REGION Network 93: Proximo Mantenimiento #1 MC060
   RUNG wire#powerrail
      { S7_Templates := "SrcType := DInt"; S7_GenerateENO := "TRUE" } Add(in1 := "Varios".UltimoMantMC060_1, in2 := "Varios".HorasMantMC060_1, out => "ProxMantMC060_1")
   END_RUNG
   // the same network as SCL:
   "ProxMantMC060_1" := "Varios".UltimoMantMC060_1 + "Varios".HorasMantMC060_1;
END_REGION

REGION Network 94: Se superaron las horas para el mantenimiento #1 MC060 / Animación Horas MAX Compresor de Alta ABC5
   RUNG wire#powerrail
      { S7_Templates := "SrcType := DInt" } GE_Contact(in1 := "HorasCmpBaja".HMMC060, in2 := "ProxMantMC060_1")
      Coil( "LimiteMantMC060_1" )
   END_RUNG
   // the same network as SCL:
   "LimiteMantMC060_1" := "HorasCmpBaja".HMMC060 >= "ProxMantMC060_1";
END_REGION

REGION Network 95: Proximo Mantenimiento #2 MC060
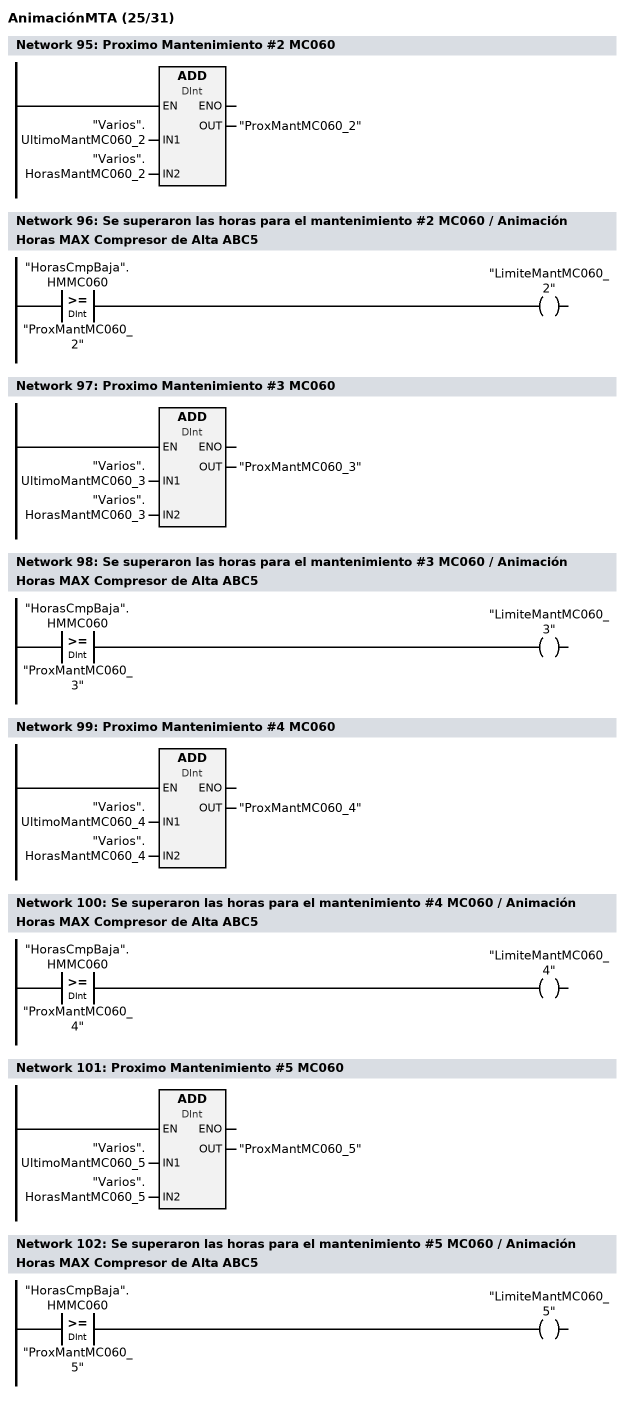
   RUNG wire#powerrail
      { S7_Templates := "SrcType := DInt"; S7_GenerateENO := "TRUE" } Add(in1 := "Varios".UltimoMantMC060_2, in2 := "Varios".HorasMantMC060_2, out => "ProxMantMC060_2")
   END_RUNG
   // the same network as SCL:
   "ProxMantMC060_2" := "Varios".UltimoMantMC060_2 + "Varios".HorasMantMC060_2;
END_REGION

REGION Network 96: Se superaron las horas para el mantenimiento #2 MC060 / Animación Horas MAX Compresor de Alta ABC5
   RUNG wire#powerrail
      { S7_Templates := "SrcType := DInt" } GE_Contact(in1 := "HorasCmpBaja".HMMC060, in2 := "ProxMantMC060_2")
      Coil( "LimiteMantMC060_2" )
   END_RUNG
   // the same network as SCL:
   "LimiteMantMC060_2" := "HorasCmpBaja".HMMC060 >= "ProxMantMC060_2";
END_REGION

REGION Network 97: Proximo Mantenimiento #3 MC060
   RUNG wire#powerrail
      { S7_Templates := "SrcType := DInt"; S7_GenerateENO := "TRUE" } Add(in1 := "Varios".UltimoMantMC060_3, in2 := "Varios".HorasMantMC060_3, out => "ProxMantMC060_3")
   END_RUNG
   // the same network as SCL:
   "ProxMantMC060_3" := "Varios".UltimoMantMC060_3 + "Varios".HorasMantMC060_3;
END_REGION

REGION Network 98: Se superaron las horas para el mantenimiento #3 MC060 / Animación Horas MAX Compresor de Alta ABC5
   RUNG wire#powerrail
      { S7_Templates := "SrcType := DInt" } GE_Contact(in1 := "HorasCmpBaja".HMMC060, in2 := "ProxMantMC060_3")
      Coil( "LimiteMantMC060_3" )
   END_RUNG
   // the same network as SCL:
   "LimiteMantMC060_3" := "HorasCmpBaja".HMMC060 >= "ProxMantMC060_3";
END_REGION

REGION Network 99: Proximo Mantenimiento #4 MC060
   RUNG wire#powerrail
      { S7_Templates := "SrcType := DInt"; S7_GenerateENO := "TRUE" } Add(in1 := "Varios".UltimoMantMC060_4, in2 := "Varios".HorasMantMC060_4, out => "ProxMantMC060_4")
   END_RUNG
   // the same network as SCL:
   "ProxMantMC060_4" := "Varios".UltimoMantMC060_4 + "Varios".HorasMantMC060_4;
END_REGION

REGION Network 100: Se superaron las horas para el mantenimiento #4 MC060 / Animación Horas MAX Compresor de Alta ABC5
   RUNG wire#powerrail
      { S7_Templates := "SrcType := DInt" } GE_Contact(in1 := "HorasCmpBaja".HMMC060, in2 := "ProxMantMC060_4")
      Coil( "LimiteMantMC060_4" )
   END_RUNG
   // the same network as SCL:
   "LimiteMantMC060_4" := "HorasCmpBaja".HMMC060 >= "ProxMantMC060_4";
END_REGION

REGION Network 101: Proximo Mantenimiento #5 MC060
   RUNG wire#powerrail
      { S7_Templates := "SrcType := DInt"; S7_GenerateENO := "TRUE" } Add(in1 := "Varios".UltimoMantMC060_5, in2 := "Varios".HorasMantMC060_5, out => "ProxMantMC060_5")
   END_RUNG
   // the same network as SCL:
   "ProxMantMC060_5" := "Varios".UltimoMantMC060_5 + "Varios".HorasMantMC060_5;
END_REGION

REGION Network 102: Se superaron las horas para el mantenimiento #5 MC060 / Animación Horas MAX Compresor de Alta ABC5
   RUNG wire#powerrail
      { S7_Templates := "SrcType := DInt" } GE_Contact(in1 := "HorasCmpBaja".HMMC060, in2 := "ProxMantMC060_5")
      Coil( "LimiteMantMC060_5" )
   END_RUNG
   // the same network as SCL:
   "LimiteMantMC060_5" := "HorasCmpBaja".HMMC060 >= "ProxMantMC060_5";
END_REGION

REGION Network 103: Proximo Mantenimiento #1 MC061
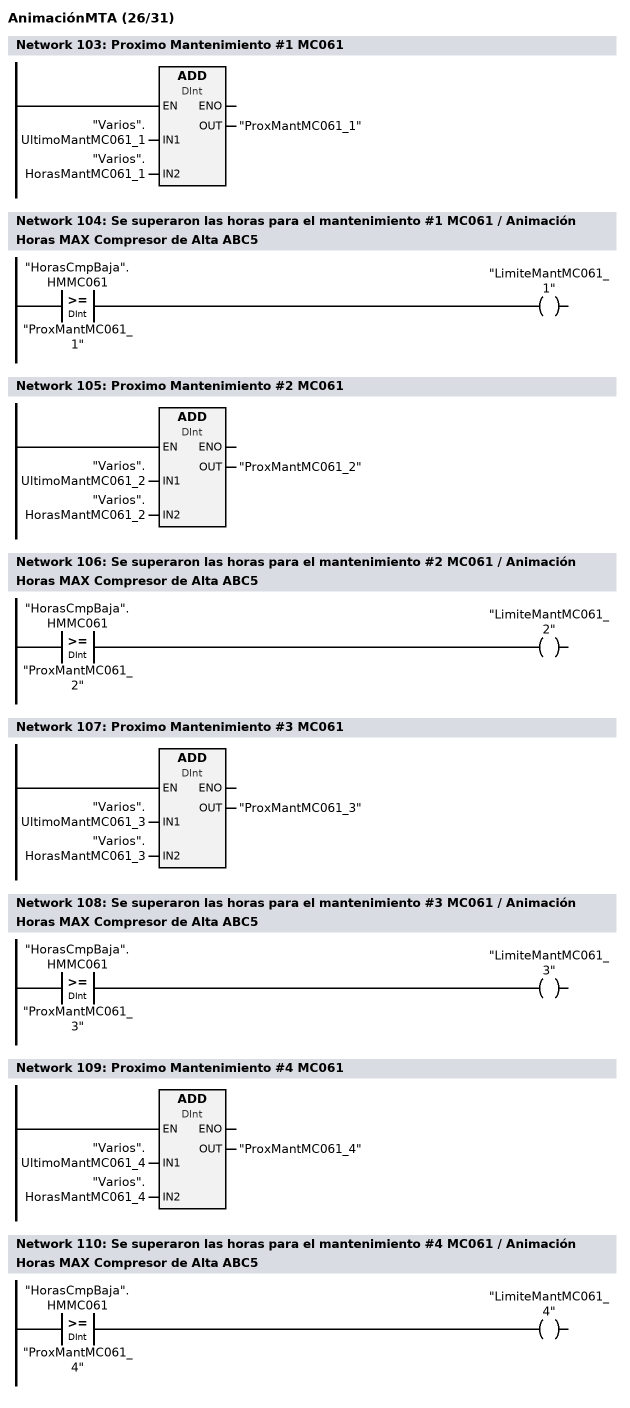
   RUNG wire#powerrail
      { S7_Templates := "SrcType := DInt"; S7_GenerateENO := "TRUE" } Add(in1 := "Varios".UltimoMantMC061_1, in2 := "Varios".HorasMantMC061_1, out => "ProxMantMC061_1")
   END_RUNG
   // the same network as SCL:
   "ProxMantMC061_1" := "Varios".UltimoMantMC061_1 + "Varios".HorasMantMC061_1;
END_REGION

REGION Network 104: Se superaron las horas para el mantenimiento #1 MC061 / Animación Horas MAX Compresor de Alta ABC5
   RUNG wire#powerrail
      { S7_Templates := "SrcType := DInt" } GE_Contact(in1 := "HorasCmpBaja".HMMC061, in2 := "ProxMantMC061_1")
      Coil( "LimiteMantMC061_1" )
   END_RUNG
   // the same network as SCL:
   "LimiteMantMC061_1" := "HorasCmpBaja".HMMC061 >= "ProxMantMC061_1";
END_REGION

REGION Network 105: Proximo Mantenimiento #2 MC061
   RUNG wire#powerrail
      { S7_Templates := "SrcType := DInt"; S7_GenerateENO := "TRUE" } Add(in1 := "Varios".UltimoMantMC061_2, in2 := "Varios".HorasMantMC061_2, out => "ProxMantMC061_2")
   END_RUNG
   // the same network as SCL:
   "ProxMantMC061_2" := "Varios".UltimoMantMC061_2 + "Varios".HorasMantMC061_2;
END_REGION

REGION Network 106: Se superaron las horas para el mantenimiento #2 MC061 / Animación Horas MAX Compresor de Alta ABC5
   RUNG wire#powerrail
      { S7_Templates := "SrcType := DInt" } GE_Contact(in1 := "HorasCmpBaja".HMMC061, in2 := "ProxMantMC061_2")
      Coil( "LimiteMantMC061_2" )
   END_RUNG
   // the same network as SCL:
   "LimiteMantMC061_2" := "HorasCmpBaja".HMMC061 >= "ProxMantMC061_2";
END_REGION

REGION Network 107: Proximo Mantenimiento #3 MC061
   RUNG wire#powerrail
      { S7_Templates := "SrcType := DInt"; S7_GenerateENO := "TRUE" } Add(in1 := "Varios".UltimoMantMC061_3, in2 := "Varios".HorasMantMC061_3, out => "ProxMantMC061_3")
   END_RUNG
   // the same network as SCL:
   "ProxMantMC061_3" := "Varios".UltimoMantMC061_3 + "Varios".HorasMantMC061_3;
END_REGION

REGION Network 108: Se superaron las horas para el mantenimiento #3 MC061 / Animación Horas MAX Compresor de Alta ABC5
   RUNG wire#powerrail
      { S7_Templates := "SrcType := DInt" } GE_Contact(in1 := "HorasCmpBaja".HMMC061, in2 := "ProxMantMC061_3")
      Coil( "LimiteMantMC061_3" )
   END_RUNG
   // the same network as SCL:
   "LimiteMantMC061_3" := "HorasCmpBaja".HMMC061 >= "ProxMantMC061_3";
END_REGION

REGION Network 109: Proximo Mantenimiento #4 MC061
   RUNG wire#powerrail
      { S7_Templates := "SrcType := DInt"; S7_GenerateENO := "TRUE" } Add(in1 := "Varios".UltimoMantMC061_4, in2 := "Varios".HorasMantMC061_4, out => "ProxMantMC061_4")
   END_RUNG
   // the same network as SCL:
   "ProxMantMC061_4" := "Varios".UltimoMantMC061_4 + "Varios".HorasMantMC061_4;
END_REGION

REGION Network 110: Se superaron las horas para el mantenimiento #4 MC061 / Animación Horas MAX Compresor de Alta ABC5
   RUNG wire#powerrail
      { S7_Templates := "SrcType := DInt" } GE_Contact(in1 := "HorasCmpBaja".HMMC061, in2 := "ProxMantMC061_4")
      Coil( "LimiteMantMC061_4" )
   END_RUNG
   // the same network as SCL:
   "LimiteMantMC061_4" := "HorasCmpBaja".HMMC061 >= "ProxMantMC061_4";
END_REGION

REGION Network 111: Proximo Mantenimiento #5 MC061
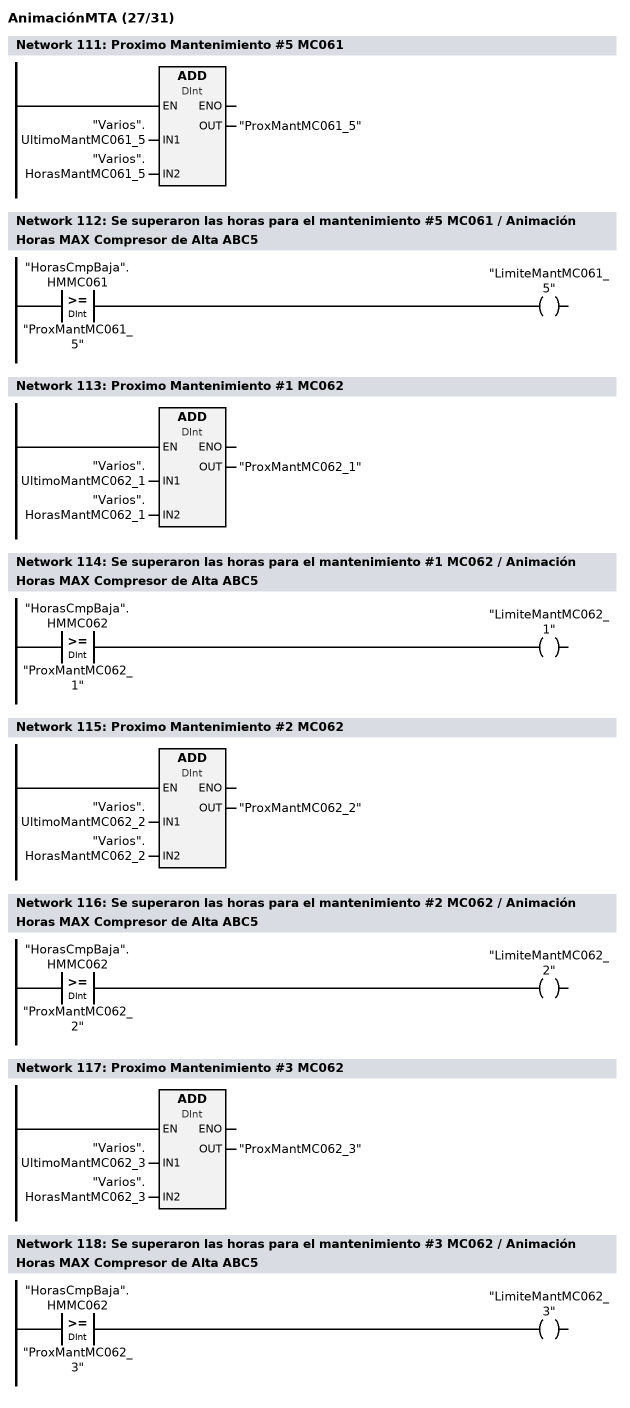
   RUNG wire#powerrail
      { S7_Templates := "SrcType := DInt"; S7_GenerateENO := "TRUE" } Add(in1 := "Varios".UltimoMantMC061_5, in2 := "Varios".HorasMantMC061_5, out => "ProxMantMC061_5")
   END_RUNG
   // the same network as SCL:
   "ProxMantMC061_5" := "Varios".UltimoMantMC061_5 + "Varios".HorasMantMC061_5;
END_REGION

REGION Network 112: Se superaron las horas para el mantenimiento #5 MC061 / Animación Horas MAX Compresor de Alta ABC5
   RUNG wire#powerrail
      { S7_Templates := "SrcType := DInt" } GE_Contact(in1 := "HorasCmpBaja".HMMC061, in2 := "ProxMantMC061_5")
      Coil( "LimiteMantMC061_5" )
   END_RUNG
   // the same network as SCL:
   "LimiteMantMC061_5" := "HorasCmpBaja".HMMC061 >= "ProxMantMC061_5";
END_REGION

REGION Network 113: Proximo Mantenimiento #1 MC062
   RUNG wire#powerrail
      { S7_Templates := "SrcType := DInt"; S7_GenerateENO := "TRUE" } Add(in1 := "Varios".UltimoMantMC062_1, in2 := "Varios".HorasMantMC062_1, out => "ProxMantMC062_1")
   END_RUNG
   // the same network as SCL:
   "ProxMantMC062_1" := "Varios".UltimoMantMC062_1 + "Varios".HorasMantMC062_1;
END_REGION

REGION Network 114: Se superaron las horas para el mantenimiento #1 MC062 / Animación Horas MAX Compresor de Alta ABC5
   RUNG wire#powerrail
      { S7_Templates := "SrcType := DInt" } GE_Contact(in1 := "HorasCmpBaja".HMMC062, in2 := "ProxMantMC062_1")
      Coil( "LimiteMantMC062_1" )
   END_RUNG
   // the same network as SCL:
   "LimiteMantMC062_1" := "HorasCmpBaja".HMMC062 >= "ProxMantMC062_1";
END_REGION

REGION Network 115: Proximo Mantenimiento #2 MC062
   RUNG wire#powerrail
      { S7_Templates := "SrcType := DInt"; S7_GenerateENO := "TRUE" } Add(in1 := "Varios".UltimoMantMC062_2, in2 := "Varios".HorasMantMC062_2, out => "ProxMantMC062_2")
   END_RUNG
   // the same network as SCL:
   "ProxMantMC062_2" := "Varios".UltimoMantMC062_2 + "Varios".HorasMantMC062_2;
END_REGION

REGION Network 116: Se superaron las horas para el mantenimiento #2 MC062 / Animación Horas MAX Compresor de Alta ABC5
   RUNG wire#powerrail
      { S7_Templates := "SrcType := DInt" } GE_Contact(in1 := "HorasCmpBaja".HMMC062, in2 := "ProxMantMC062_2")
      Coil( "LimiteMantMC062_2" )
   END_RUNG
   // the same network as SCL:
   "LimiteMantMC062_2" := "HorasCmpBaja".HMMC062 >= "ProxMantMC062_2";
END_REGION

REGION Network 117: Proximo Mantenimiento #3 MC062
   RUNG wire#powerrail
      { S7_Templates := "SrcType := DInt"; S7_GenerateENO := "TRUE" } Add(in1 := "Varios".UltimoMantMC062_3, in2 := "Varios".HorasMantMC062_3, out => "ProxMantMC062_3")
   END_RUNG
   // the same network as SCL:
   "ProxMantMC062_3" := "Varios".UltimoMantMC062_3 + "Varios".HorasMantMC062_3;
END_REGION

REGION Network 118: Se superaron las horas para el mantenimiento #3 MC062 / Animación Horas MAX Compresor de Alta ABC5
   RUNG wire#powerrail
      { S7_Templates := "SrcType := DInt" } GE_Contact(in1 := "HorasCmpBaja".HMMC062, in2 := "ProxMantMC062_3")
      Coil( "LimiteMantMC062_3" )
   END_RUNG
   // the same network as SCL:
   "LimiteMantMC062_3" := "HorasCmpBaja".HMMC062 >= "ProxMantMC062_3";
END_REGION

REGION Network 119: Proximo Mantenimiento #4 MC062
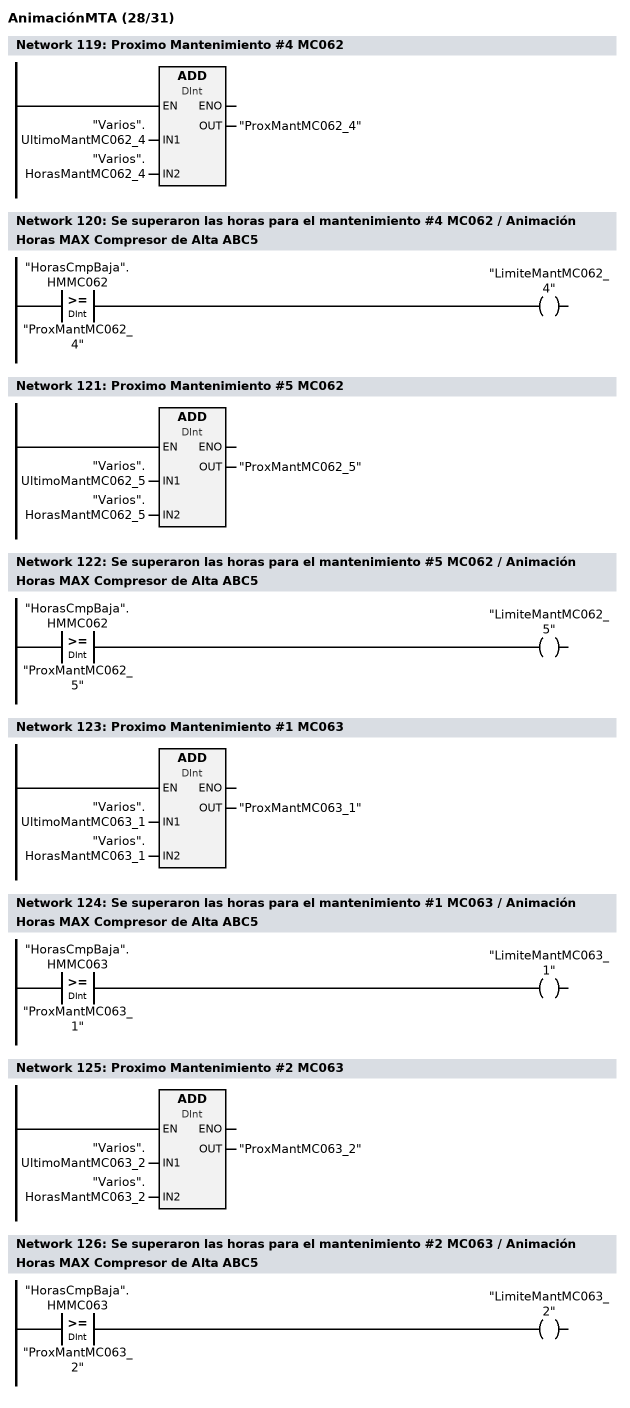
   RUNG wire#powerrail
      { S7_Templates := "SrcType := DInt"; S7_GenerateENO := "TRUE" } Add(in1 := "Varios".UltimoMantMC062_4, in2 := "Varios".HorasMantMC062_4, out => "ProxMantMC062_4")
   END_RUNG
   // the same network as SCL:
   "ProxMantMC062_4" := "Varios".UltimoMantMC062_4 + "Varios".HorasMantMC062_4;
END_REGION

REGION Network 120: Se superaron las horas para el mantenimiento #4 MC062 / Animación Horas MAX Compresor de Alta ABC5
   RUNG wire#powerrail
      { S7_Templates := "SrcType := DInt" } GE_Contact(in1 := "HorasCmpBaja".HMMC062, in2 := "ProxMantMC062_4")
      Coil( "LimiteMantMC062_4" )
   END_RUNG
   // the same network as SCL:
   "LimiteMantMC062_4" := "HorasCmpBaja".HMMC062 >= "ProxMantMC062_4";
END_REGION

REGION Network 121: Proximo Mantenimiento #5 MC062
   RUNG wire#powerrail
      { S7_Templates := "SrcType := DInt"; S7_GenerateENO := "TRUE" } Add(in1 := "Varios".UltimoMantMC062_5, in2 := "Varios".HorasMantMC062_5, out => "ProxMantMC062_5")
   END_RUNG
   // the same network as SCL:
   "ProxMantMC062_5" := "Varios".UltimoMantMC062_5 + "Varios".HorasMantMC062_5;
END_REGION

REGION Network 122: Se superaron las horas para el mantenimiento #5 MC062 / Animación Horas MAX Compresor de Alta ABC5
   RUNG wire#powerrail
      { S7_Templates := "SrcType := DInt" } GE_Contact(in1 := "HorasCmpBaja".HMMC062, in2 := "ProxMantMC062_5")
      Coil( "LimiteMantMC062_5" )
   END_RUNG
   // the same network as SCL:
   "LimiteMantMC062_5" := "HorasCmpBaja".HMMC062 >= "ProxMantMC062_5";
END_REGION

REGION Network 123: Proximo Mantenimiento #1 MC063
   RUNG wire#powerrail
      { S7_Templates := "SrcType := DInt"; S7_GenerateENO := "TRUE" } Add(in1 := "Varios".UltimoMantMC063_1, in2 := "Varios".HorasMantMC063_1, out => "ProxMantMC063_1")
   END_RUNG
   // the same network as SCL:
   "ProxMantMC063_1" := "Varios".UltimoMantMC063_1 + "Varios".HorasMantMC063_1;
END_REGION

REGION Network 124: Se superaron las horas para el mantenimiento #1 MC063 / Animación Horas MAX Compresor de Alta ABC5
   RUNG wire#powerrail
      { S7_Templates := "SrcType := DInt" } GE_Contact(in1 := "HorasCmpBaja".HMMC063, in2 := "ProxMantMC063_1")
      Coil( "LimiteMantMC063_1" )
   END_RUNG
   // the same network as SCL:
   "LimiteMantMC063_1" := "HorasCmpBaja".HMMC063 >= "ProxMantMC063_1";
END_REGION

REGION Network 125: Proximo Mantenimiento #2 MC063
   RUNG wire#powerrail
      { S7_Templates := "SrcType := DInt"; S7_GenerateENO := "TRUE" } Add(in1 := "Varios".UltimoMantMC063_2, in2 := "Varios".HorasMantMC063_2, out => "ProxMantMC063_2")
   END_RUNG
   // the same network as SCL:
   "ProxMantMC063_2" := "Varios".UltimoMantMC063_2 + "Varios".HorasMantMC063_2;
END_REGION

REGION Network 126: Se superaron las horas para el mantenimiento #2 MC063 / Animación Horas MAX Compresor de Alta ABC5
   RUNG wire#powerrail
      { S7_Templates := "SrcType := DInt" } GE_Contact(in1 := "HorasCmpBaja".HMMC063, in2 := "ProxMantMC063_2")
      Coil( "LimiteMantMC063_2" )
   END_RUNG
   // the same network as SCL:
   "LimiteMantMC063_2" := "HorasCmpBaja".HMMC063 >= "ProxMantMC063_2";
END_REGION

REGION Network 127: Proximo Mantenimiento #3 MC063
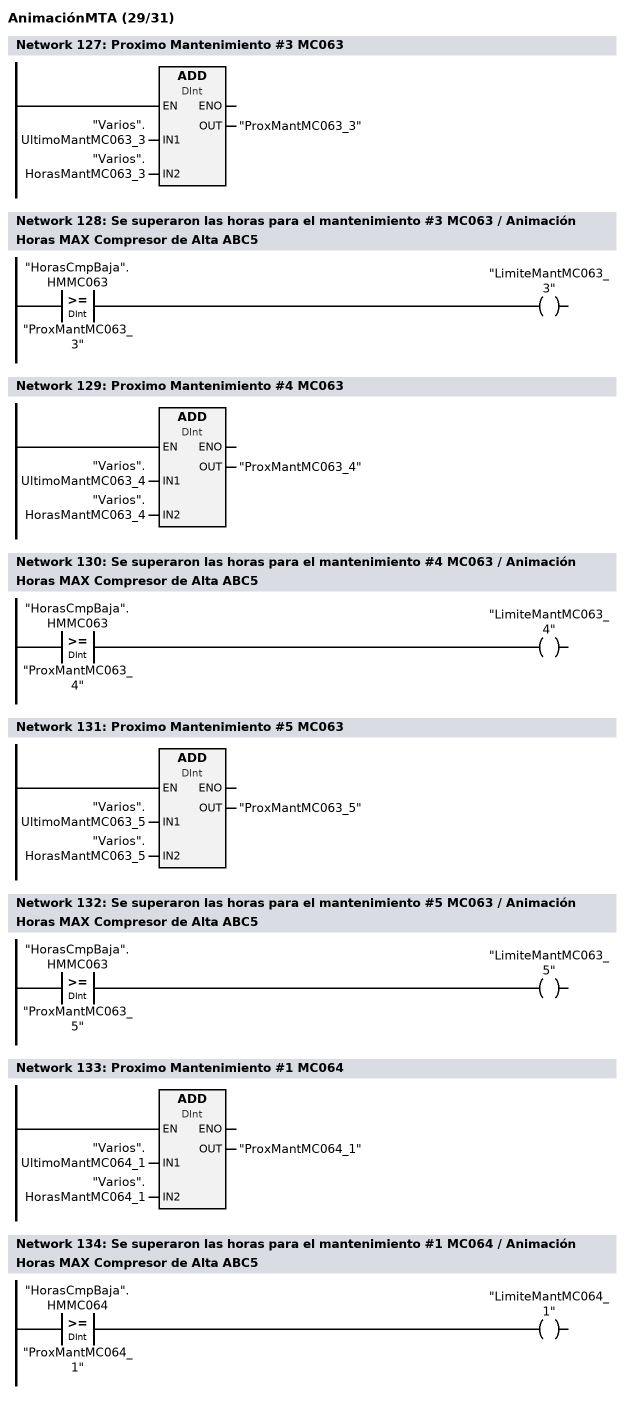
   RUNG wire#powerrail
      { S7_Templates := "SrcType := DInt"; S7_GenerateENO := "TRUE" } Add(in1 := "Varios".UltimoMantMC063_3, in2 := "Varios".HorasMantMC063_3, out => "ProxMantMC063_3")
   END_RUNG
   // the same network as SCL:
   "ProxMantMC063_3" := "Varios".UltimoMantMC063_3 + "Varios".HorasMantMC063_3;
END_REGION

REGION Network 128: Se superaron las horas para el mantenimiento #3 MC063 / Animación Horas MAX Compresor de Alta ABC5
   RUNG wire#powerrail
      { S7_Templates := "SrcType := DInt" } GE_Contact(in1 := "HorasCmpBaja".HMMC063, in2 := "ProxMantMC063_3")
      Coil( "LimiteMantMC063_3" )
   END_RUNG
   // the same network as SCL:
   "LimiteMantMC063_3" := "HorasCmpBaja".HMMC063 >= "ProxMantMC063_3";
END_REGION

REGION Network 129: Proximo Mantenimiento #4 MC063
   RUNG wire#powerrail
      { S7_Templates := "SrcType := DInt"; S7_GenerateENO := "TRUE" } Add(in1 := "Varios".UltimoMantMC063_4, in2 := "Varios".HorasMantMC063_4, out => "ProxMantMC063_4")
   END_RUNG
   // the same network as SCL:
   "ProxMantMC063_4" := "Varios".UltimoMantMC063_4 + "Varios".HorasMantMC063_4;
END_REGION

REGION Network 130: Se superaron las horas para el mantenimiento #4 MC063 / Animación Horas MAX Compresor de Alta ABC5
   RUNG wire#powerrail
      { S7_Templates := "SrcType := DInt" } GE_Contact(in1 := "HorasCmpBaja".HMMC063, in2 := "ProxMantMC063_4")
      Coil( "LimiteMantMC063_4" )
   END_RUNG
   // the same network as SCL:
   "LimiteMantMC063_4" := "HorasCmpBaja".HMMC063 >= "ProxMantMC063_4";
END_REGION

REGION Network 131: Proximo Mantenimiento #5 MC063
   RUNG wire#powerrail
      { S7_Templates := "SrcType := DInt"; S7_GenerateENO := "TRUE" } Add(in1 := "Varios".UltimoMantMC063_5, in2 := "Varios".HorasMantMC063_5, out => "ProxMantMC063_5")
   END_RUNG
   // the same network as SCL:
   "ProxMantMC063_5" := "Varios".UltimoMantMC063_5 + "Varios".HorasMantMC063_5;
END_REGION

REGION Network 132: Se superaron las horas para el mantenimiento #5 MC063 / Animación Horas MAX Compresor de Alta ABC5
   RUNG wire#powerrail
      { S7_Templates := "SrcType := DInt" } GE_Contact(in1 := "HorasCmpBaja".HMMC063, in2 := "ProxMantMC063_5")
      Coil( "LimiteMantMC063_5" )
   END_RUNG
   // the same network as SCL:
   "LimiteMantMC063_5" := "HorasCmpBaja".HMMC063 >= "ProxMantMC063_5";
END_REGION

REGION Network 133: Proximo Mantenimiento #1 MC064
   RUNG wire#powerrail
      { S7_Templates := "SrcType := DInt"; S7_GenerateENO := "TRUE" } Add(in1 := "Varios".UltimoMantMC064_1, in2 := "Varios".HorasMantMC064_1, out => "ProxMantMC064_1")
   END_RUNG
   // the same network as SCL:
   "ProxMantMC064_1" := "Varios".UltimoMantMC064_1 + "Varios".HorasMantMC064_1;
END_REGION

REGION Network 134: Se superaron las horas para el mantenimiento #1 MC064 / Animación Horas MAX Compresor de Alta ABC5
   RUNG wire#powerrail
      { S7_Templates := "SrcType := DInt" } GE_Contact(in1 := "HorasCmpBaja".HMMC064, in2 := "ProxMantMC064_1")
      Coil( "LimiteMantMC064_1" )
   END_RUNG
   // the same network as SCL:
   "LimiteMantMC064_1" := "HorasCmpBaja".HMMC064 >= "ProxMantMC064_1";
END_REGION

REGION Network 135: Proximo Mantenimiento #2 MC064
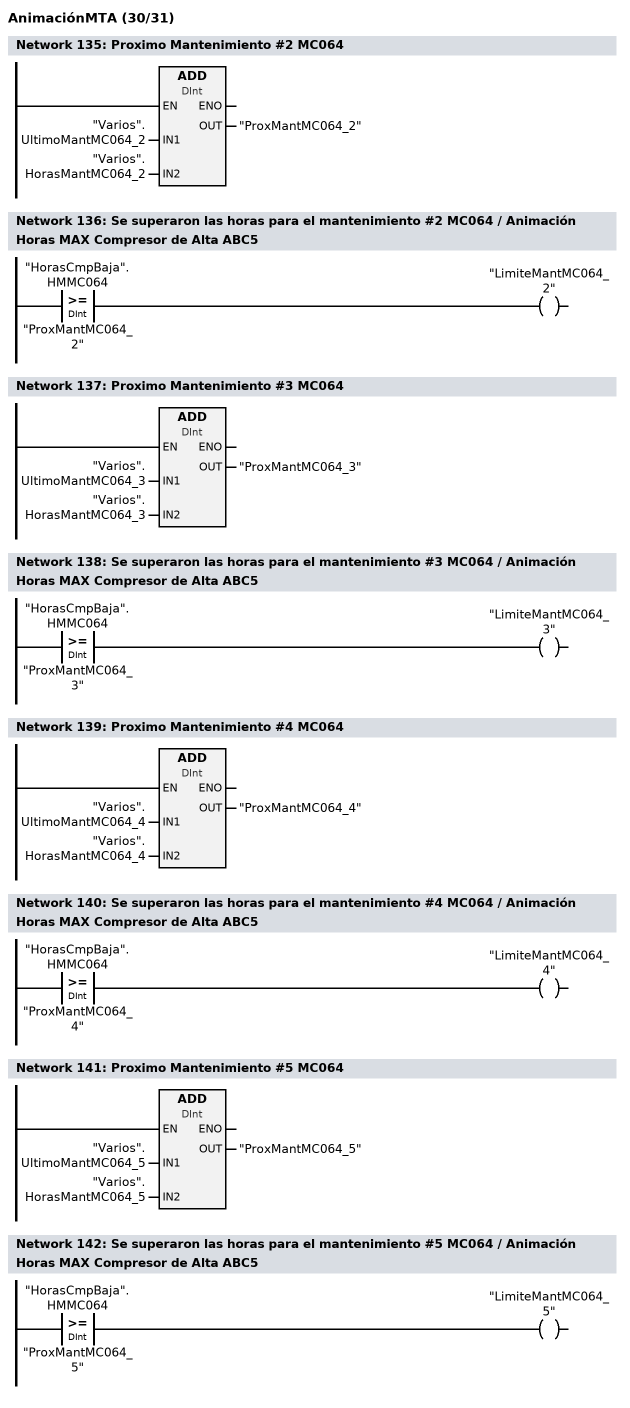
   RUNG wire#powerrail
      { S7_Templates := "SrcType := DInt"; S7_GenerateENO := "TRUE" } Add(in1 := "Varios".UltimoMantMC064_2, in2 := "Varios".HorasMantMC064_2, out => "ProxMantMC064_2")
   END_RUNG
   // the same network as SCL:
   "ProxMantMC064_2" := "Varios".UltimoMantMC064_2 + "Varios".HorasMantMC064_2;
END_REGION

REGION Network 136: Se superaron las horas para el mantenimiento #2 MC064 / Animación Horas MAX Compresor de Alta ABC5
   RUNG wire#powerrail
      { S7_Templates := "SrcType := DInt" } GE_Contact(in1 := "HorasCmpBaja".HMMC064, in2 := "ProxMantMC064_2")
      Coil( "LimiteMantMC064_2" )
   END_RUNG
   // the same network as SCL:
   "LimiteMantMC064_2" := "HorasCmpBaja".HMMC064 >= "ProxMantMC064_2";
END_REGION

REGION Network 137: Proximo Mantenimiento #3 MC064
   RUNG wire#powerrail
      { S7_Templates := "SrcType := DInt"; S7_GenerateENO := "TRUE" } Add(in1 := "Varios".UltimoMantMC064_3, in2 := "Varios".HorasMantMC064_3, out => "ProxMantMC064_3")
   END_RUNG
   // the same network as SCL:
   "ProxMantMC064_3" := "Varios".UltimoMantMC064_3 + "Varios".HorasMantMC064_3;
END_REGION

REGION Network 138: Se superaron las horas para el mantenimiento #3 MC064 / Animación Horas MAX Compresor de Alta ABC5
   RUNG wire#powerrail
      { S7_Templates := "SrcType := DInt" } GE_Contact(in1 := "HorasCmpBaja".HMMC064, in2 := "ProxMantMC064_3")
      Coil( "LimiteMantMC064_3" )
   END_RUNG
   // the same network as SCL:
   "LimiteMantMC064_3" := "HorasCmpBaja".HMMC064 >= "ProxMantMC064_3";
END_REGION

REGION Network 139: Proximo Mantenimiento #4 MC064
   RUNG wire#powerrail
      { S7_Templates := "SrcType := DInt"; S7_GenerateENO := "TRUE" } Add(in1 := "Varios".UltimoMantMC064_4, in2 := "Varios".HorasMantMC064_4, out => "ProxMantMC064_4")
   END_RUNG
   // the same network as SCL:
   "ProxMantMC064_4" := "Varios".UltimoMantMC064_4 + "Varios".HorasMantMC064_4;
END_REGION

REGION Network 140: Se superaron las horas para el mantenimiento #4 MC064 / Animación Horas MAX Compresor de Alta ABC5
   RUNG wire#powerrail
      { S7_Templates := "SrcType := DInt" } GE_Contact(in1 := "HorasCmpBaja".HMMC064, in2 := "ProxMantMC064_4")
      Coil( "LimiteMantMC064_4" )
   END_RUNG
   // the same network as SCL:
   "LimiteMantMC064_4" := "HorasCmpBaja".HMMC064 >= "ProxMantMC064_4";
END_REGION

REGION Network 141: Proximo Mantenimiento #5 MC064
   RUNG wire#powerrail
      { S7_Templates := "SrcType := DInt"; S7_GenerateENO := "TRUE" } Add(in1 := "Varios".UltimoMantMC064_5, in2 := "Varios".HorasMantMC064_5, out => "ProxMantMC064_5")
   END_RUNG
   // the same network as SCL:
   "ProxMantMC064_5" := "Varios".UltimoMantMC064_5 + "Varios".HorasMantMC064_5;
END_REGION

REGION Network 142: Se superaron las horas para el mantenimiento #5 MC064 / Animación Horas MAX Compresor de Alta ABC5
   RUNG wire#powerrail
      { S7_Templates := "SrcType := DInt" } GE_Contact(in1 := "HorasCmpBaja".HMMC064, in2 := "ProxMantMC064_5")
      Coil( "LimiteMantMC064_5" )
   END_RUNG
   // the same network as SCL:
   "LimiteMantMC064_5" := "HorasCmpBaja".HMMC064 >= "ProxMantMC064_5";
END_REGION

REGION Network 143: Próximo Mantenimento Booster 1
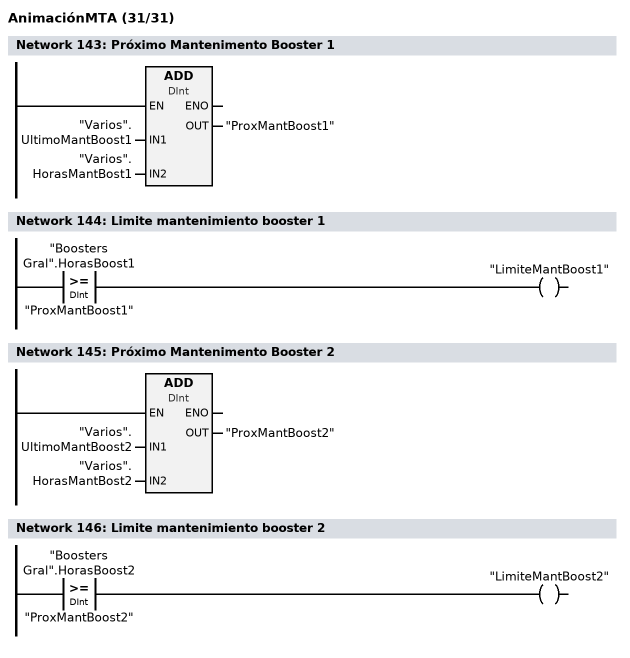
   RUNG wire#powerrail
      { S7_Templates := "SrcType := DInt"; S7_GenerateENO := "TRUE" } Add(in1 := "Varios".UltimoMantBoost1, in2 := "Varios".HorasMantBost1, out => "ProxMantBoost1")
   END_RUNG
   // the same network as SCL:
   "ProxMantBoost1" := "Varios".UltimoMantBoost1 + "Varios".HorasMantBost1;
END_REGION

REGION Network 144: Limite mantenimiento booster 1
   RUNG wire#powerrail
      { S7_Templates := "SrcType := DInt" } GE_Contact(in1 := "Boosters Gral".HorasBoost1, in2 := "ProxMantBoost1")
      Coil( "LimiteMantBoost1" )
   END_RUNG
   // the same network as SCL:
   "LimiteMantBoost1" := "Boosters Gral".HorasBoost1 >= "ProxMantBoost1";
END_REGION

REGION Network 145: Próximo Mantenimento Booster 2
   RUNG wire#powerrail
      { S7_Templates := "SrcType := DInt"; S7_GenerateENO := "TRUE" } Add(in1 := "Varios".UltimoMantBoost2, in2 := "Varios".HorasMantBost2, out => "ProxMantBoost2")
   END_RUNG
   // the same network as SCL:
   "ProxMantBoost2" := "Varios".UltimoMantBoost2 + "Varios".HorasMantBost2;
END_REGION

REGION Network 146: Limite mantenimiento booster 2
   RUNG wire#powerrail
      { S7_Templates := "SrcType := DInt" } GE_Contact(in1 := "Boosters Gral".HorasBoost2, in2 := "ProxMantBoost2")
      Coil( "LimiteMantBoost2" )
   END_RUNG
   // the same network as SCL:
   "LimiteMantBoost2" := "Boosters Gral".HorasBoost2 >= "ProxMantBoost2";
END_REGION
END_FUNCTION

FUNCTION "Motores-PanelMTA" : Void   // FC3, LAD
{ S7_Optimized_Access := 'FALSE' }
VERSION : 0.1
BEGIN

REGION Network 1: Comandos desde Panel para MP010 - Bomba Principal Ch. Soplado
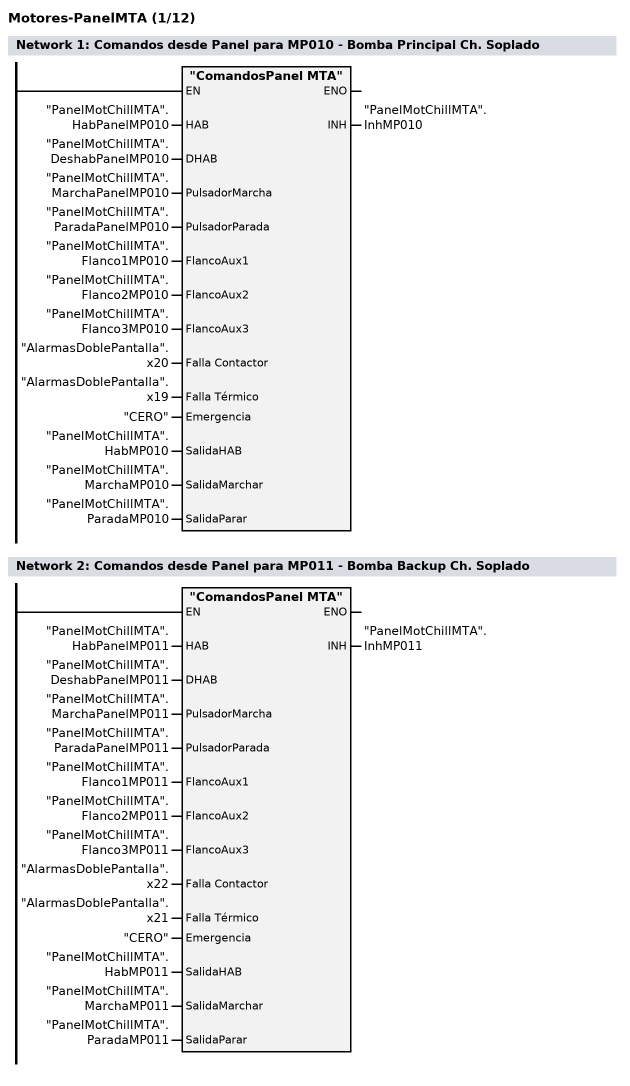
   RUNG wire#powerrail
      "ComandosPanel MTA"(HAB := "PanelMotChillMTA".HabPanelMP010, DHAB := "PanelMotChillMTA".DeshabPanelMP010, PulsadorMarcha := "PanelMotChillMTA".MarchaPanelMP010, PulsadorParada := "PanelMotChillMTA".ParadaPanelMP010, FlancoAux1 := "PanelMotChillMTA".Flanco1MP010, FlancoAux2 := "PanelMotChillMTA".Flanco2MP010, FlancoAux3 := "PanelMotChillMTA".Flanco3MP010, "Falla Contactor" := "AlarmasDoblePantalla".x20, "Falla Térmico" := "AlarmasDoblePantalla".x19, Emergencia := "CERO", INH => "PanelMotChillMTA".InhMP010, SalidaHAB := "PanelMotChillMTA".HabMP010, SalidaMarchar := "PanelMotChillMTA".MarchaMP010, SalidaParar := "PanelMotChillMTA".ParadaMP010)
   END_RUNG
   // the same network as SCL:
   "ComandosPanel MTA"(HAB := "PanelMotChillMTA".HabPanelMP010,
                       DHAB := "PanelMotChillMTA".DeshabPanelMP010,
                       PulsadorMarcha := "PanelMotChillMTA".MarchaPanelMP010,
                       PulsadorParada := "PanelMotChillMTA".ParadaPanelMP010,
                       FlancoAux1 := "PanelMotChillMTA".Flanco1MP010,
                       FlancoAux2 := "PanelMotChillMTA".Flanco2MP010,
                       FlancoAux3 := "PanelMotChillMTA".Flanco3MP010,
                       "Falla Contactor" := "AlarmasDoblePantalla".x20,
                       "Falla Térmico" := "AlarmasDoblePantalla".x19,
                       Emergencia := "CERO",
                       SalidaHAB := "PanelMotChillMTA".HabMP010,
                       SalidaMarchar := "PanelMotChillMTA".MarchaMP010,
                       SalidaParar := "PanelMotChillMTA".ParadaMP010,
                       INH => "PanelMotChillMTA".InhMP010);
END_REGION

REGION Network 2: Comandos desde Panel para MP011 - Bomba Backup Ch. Soplado
   RUNG wire#powerrail
      "ComandosPanel MTA"(HAB := "PanelMotChillMTA".HabPanelMP011, DHAB := "PanelMotChillMTA".DeshabPanelMP011, PulsadorMarcha := "PanelMotChillMTA".MarchaPanelMP011, PulsadorParada := "PanelMotChillMTA".ParadaPanelMP011, FlancoAux1 := "PanelMotChillMTA".Flanco1MP011, FlancoAux2 := "PanelMotChillMTA".Flanco2MP011, FlancoAux3 := "PanelMotChillMTA".Flanco3MP011, "Falla Contactor" := "AlarmasDoblePantalla".x22, "Falla Térmico" := "AlarmasDoblePantalla".x21, Emergencia := "CERO", INH => "PanelMotChillMTA".InhMP011, SalidaHAB := "PanelMotChillMTA".HabMP011, SalidaMarchar := "PanelMotChillMTA".MarchaMP011, SalidaParar := "PanelMotChillMTA".ParadaMP011)
   END_RUNG
   // the same network as SCL:
   "ComandosPanel MTA"(HAB := "PanelMotChillMTA".HabPanelMP011,
                       DHAB := "PanelMotChillMTA".DeshabPanelMP011,
                       PulsadorMarcha := "PanelMotChillMTA".MarchaPanelMP011,
                       PulsadorParada := "PanelMotChillMTA".ParadaPanelMP011,
                       FlancoAux1 := "PanelMotChillMTA".Flanco1MP011,
                       FlancoAux2 := "PanelMotChillMTA".Flanco2MP011,
                       FlancoAux3 := "PanelMotChillMTA".Flanco3MP011,
                       "Falla Contactor" := "AlarmasDoblePantalla".x22,
                       "Falla Térmico" := "AlarmasDoblePantalla".x21,
                       Emergencia := "CERO",
                       SalidaHAB := "PanelMotChillMTA".HabMP011,
                       SalidaMarchar := "PanelMotChillMTA".MarchaMP011,
                       SalidaParar := "PanelMotChillMTA".ParadaMP011,
                       INH => "PanelMotChillMTA".InhMP011);
END_REGION

REGION Network 3: Comandos desde Panel para MP012 - Bomba Principal Ch. Envasado
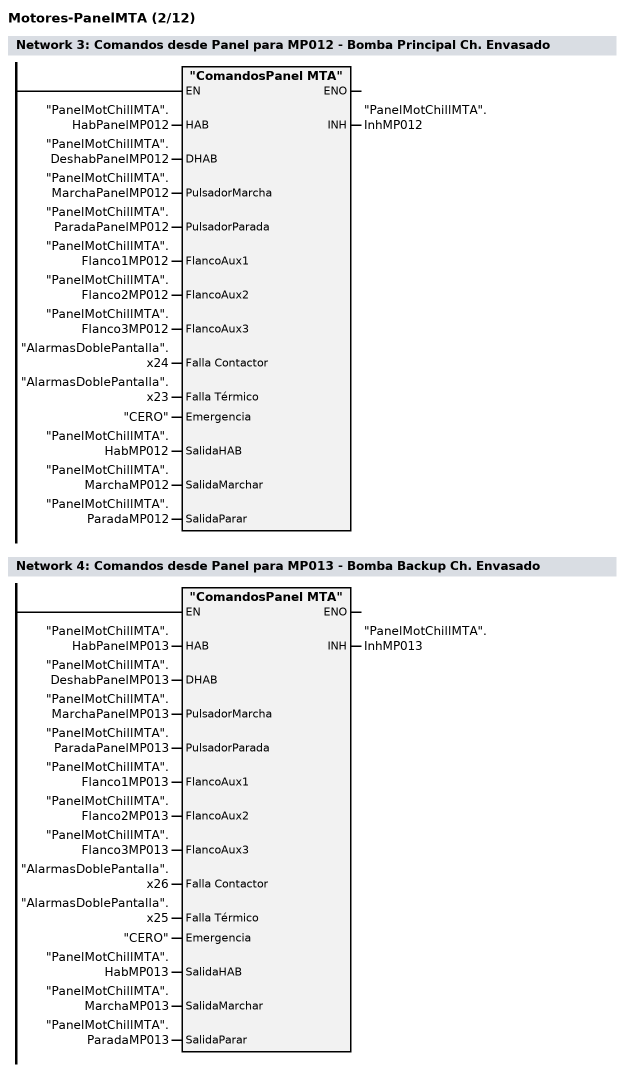
   RUNG wire#powerrail
      "ComandosPanel MTA"(HAB := "PanelMotChillMTA".HabPanelMP012, DHAB := "PanelMotChillMTA".DeshabPanelMP012, PulsadorMarcha := "PanelMotChillMTA".MarchaPanelMP012, PulsadorParada := "PanelMotChillMTA".ParadaPanelMP012, FlancoAux1 := "PanelMotChillMTA".Flanco1MP012, FlancoAux2 := "PanelMotChillMTA".Flanco2MP012, FlancoAux3 := "PanelMotChillMTA".Flanco3MP012, "Falla Contactor" := "AlarmasDoblePantalla".x24, "Falla Térmico" := "AlarmasDoblePantalla".x23, Emergencia := "CERO", INH => "PanelMotChillMTA".InhMP012, SalidaHAB := "PanelMotChillMTA".HabMP012, SalidaMarchar := "PanelMotChillMTA".MarchaMP012, SalidaParar := "PanelMotChillMTA".ParadaMP012)
   END_RUNG
   // the same network as SCL:
   "ComandosPanel MTA"(HAB := "PanelMotChillMTA".HabPanelMP012,
                       DHAB := "PanelMotChillMTA".DeshabPanelMP012,
                       PulsadorMarcha := "PanelMotChillMTA".MarchaPanelMP012,
                       PulsadorParada := "PanelMotChillMTA".ParadaPanelMP012,
                       FlancoAux1 := "PanelMotChillMTA".Flanco1MP012,
                       FlancoAux2 := "PanelMotChillMTA".Flanco2MP012,
                       FlancoAux3 := "PanelMotChillMTA".Flanco3MP012,
                       "Falla Contactor" := "AlarmasDoblePantalla".x24,
                       "Falla Térmico" := "AlarmasDoblePantalla".x23,
                       Emergencia := "CERO",
                       SalidaHAB := "PanelMotChillMTA".HabMP012,
                       SalidaMarchar := "PanelMotChillMTA".MarchaMP012,
                       SalidaParar := "PanelMotChillMTA".ParadaMP012,
                       INH => "PanelMotChillMTA".InhMP012);
END_REGION

REGION Network 4: Comandos desde Panel para MP013 - Bomba Backup Ch. Envasado
   RUNG wire#powerrail
      "ComandosPanel MTA"(HAB := "PanelMotChillMTA".HabPanelMP013, DHAB := "PanelMotChillMTA".DeshabPanelMP013, PulsadorMarcha := "PanelMotChillMTA".MarchaPanelMP013, PulsadorParada := "PanelMotChillMTA".ParadaPanelMP013, FlancoAux1 := "PanelMotChillMTA".Flanco1MP013, FlancoAux2 := "PanelMotChillMTA".Flanco2MP013, FlancoAux3 := "PanelMotChillMTA".Flanco3MP013, "Falla Contactor" := "AlarmasDoblePantalla".x26, "Falla Térmico" := "AlarmasDoblePantalla".x25, Emergencia := "CERO", INH => "PanelMotChillMTA".InhMP013, SalidaHAB := "PanelMotChillMTA".HabMP013, SalidaMarchar := "PanelMotChillMTA".MarchaMP013, SalidaParar := "PanelMotChillMTA".ParadaMP013)
   END_RUNG
   // the same network as SCL:
   "ComandosPanel MTA"(HAB := "PanelMotChillMTA".HabPanelMP013,
                       DHAB := "PanelMotChillMTA".DeshabPanelMP013,
                       PulsadorMarcha := "PanelMotChillMTA".MarchaPanelMP013,
                       PulsadorParada := "PanelMotChillMTA".ParadaPanelMP013,
                       FlancoAux1 := "PanelMotChillMTA".Flanco1MP013,
                       FlancoAux2 := "PanelMotChillMTA".Flanco2MP013,
                       FlancoAux3 := "PanelMotChillMTA".Flanco3MP013,
                       "Falla Contactor" := "AlarmasDoblePantalla".x26,
                       "Falla Térmico" := "AlarmasDoblePantalla".x25,
                       Emergencia := "CERO",
                       SalidaHAB := "PanelMotChillMTA".HabMP013,
                       SalidaMarchar := "PanelMotChillMTA".MarchaMP013,
                       SalidaParar := "PanelMotChillMTA".ParadaMP013,
                       INH => "PanelMotChillMTA".InhMP013);
END_REGION

REGION Network 5: Comandos desde Panel para MP018 - Bomba 1 Torres de enfriamiento Chillers
